screen "eProC - Edición Recetas" 1280x770, template "Template"
   RecipeView "Visor de recetas_1" at 25,54 size 1221x597; Recipe "Pieza"
   TextField "Campo de texto_2" at 43,32 size 125x22; Text 'Edición de Recetas'
   Button "Template_Plantilla_Bouton_12" at 937,715 size 150x53; TextOff 'Ajustes Avanzados SYSTEM'; Authorization "Nivel 2"
      on Press: ActivateScreen("eProC - Avanzado", 0)
   Button "Template_Plantilla_Botón_2" at 128,688 size 150x29; TextOff 'EDICIÓN RECETAS'
   Button "Template_Plantilla_Botón_3" at 129,715 size 150x53; TextOff 'SELECCIÓN RECETAS'
      on Click: ActivateScreen("eProC - Recetas", 0)

screen "HabAlarmas5" 1280x770, template "Template"
   TextField "Campo de texto_1" at 117,85 size 297x18; Text '057 - Falla en Plegador 1 al intentar desactivar fijación'
   TextField "Campo de texto_2" at 117,129 size 357x18; Text '058 - Falla en Plegador 1 al intentar desactivar orden de plegado'
   TextField "Campo de texto_3" at 117,173 size 267x18; Text '059 - Falla en Plegador 1 al intentar subir prensa'
   TextField "Campo de texto_4" at 117,217 size 387x18; Text '060 - Falla en Plegador 1 al intentar bajar primera extensión de prensa'
   TextField "Campo de texto_5" at 117,261 size 297x18; Text '061 - Falla en Plegador 2 al intentar desactivar fijación'
   TextField "Campo de texto_6g" at 117,305 size 357x18; Text '062 - Falla en Plegador 2 al intentar desactivar orden de plegado'
   TextField "Campo de texto_7" at 117,349 size 267x18; Text '063 - Falla en Plegador 2 al intentar subir prensa'
   TextField "Campo de texto_8" at 117,393 size 386x18; Text '064 - Falla en Plegador 2 al intentar subir primera extensión de prensa'
   TextField "Campo de texto_9" at 117,437 size 216x18; Text '065 - Falla al transladar Araña (Avance)'
   TextField "Campo de texto_10" at 117,483 size 135x18; Text '066 - Falla al subir Araña'
   TextField "Campo de texto_11" at 117,525 size 136x18; Text '067 - Falla al bajar Araña'
   TextField "Campo de texto_12" at 117,571 size 135x18; Text '068 - Falla al subir Araña'
   TextField "Campo de texto_13" at 117,613 size 37x18; Text '069 -'
   TextField "Campo de texto_14" at 117,657 size 37x18; Text '070 -'
   Switch "Interruptor_1" at 48,77 size 59x33; TextOff 'SI'; TextOn 'NO'; CaptionText 'Switch'; PictureOff "Check"; PictureOn "UnCheck"
      ProcessValue <- "Desactivar_Falla57"
   Switch "Interruptor_2" at 48,121 size 59x33; TextOff 'SI'; TextOn 'NO'; CaptionText 'Switch'; PictureOff "Check"; PictureOn "UnCheck"
      ProcessValue <- "Desactivar_Falla58"
   Switch "Interruptor_3" at 48,165 size 59x33; TextOff 'SI'; TextOn 'NO'; CaptionText 'Switch'; PictureOff "Check"; PictureOn "UnCheck"
      ProcessValue <- "Desactivar_Falla59"
   Switch "Interruptor_4" at 48,209 size 59x33; TextOff 'SI'; TextOn 'NO'; CaptionText 'Switch'; PictureOff "Check"; PictureOn "UnCheck"
      ProcessValue <- "Desactivar_Falla60"
   Switch "Interruptor_5" at 48,253 size 59x33; TextOff 'SI'; TextOn 'NO'; CaptionText 'Switch'; PictureOff "Check"; PictureOn "UnCheck"
      ProcessValue <- "Desactivar_Falla61"
   Switch "Interruptor_6" at 48,297 size 59x33; TextOff 'SI'; TextOn 'NO'; CaptionText 'Switch'; PictureOff "Check"; PictureOn "UnCheck"
      ProcessValue <- "Desactivar_Falla62"
   Switch "Interruptor_7" at 48,341 size 59x33; TextOff 'SI'; TextOn 'NO'; CaptionText 'Switch'; PictureOff "Check"; PictureOn "UnCheck"
      ProcessValue <- "Desactivar_Falla63"
   Switch "Interruptor_8" at 48,385 size 59x33; TextOff 'SI'; TextOn 'NO'; CaptionText 'Switch'; PictureOff "Check"; PictureOn "UnCheck"
      ProcessValue <- "Desactivar_Falla64"
   Switch "Interruptor_9" at 48,429 size 59x33; TextOff 'SI'; TextOn 'NO'; CaptionText 'Switch'; PictureOff "Check"; PictureOn "UnCheck"
      ProcessValue <- "Desactivar_Falla65"
   Switch "Interruptor_10" at 48,473 size 59x33; TextOff 'SI'; TextOn 'NO'; CaptionText 'Switch'; PictureOff "Check"; PictureOn "UnCheck"
      ProcessValue <- "Desactivar_Falla66"
   Switch "Interruptor_11" at 48,517 size 59x33; TextOff 'SI'; TextOn 'NO'; CaptionText 'Switch'; PictureOff "Check"; PictureOn "UnCheck"
      ProcessValue <- "Desactivar_Falla67"
   Switch "Interruptor_12" at 48,561 size 59x33; TextOff 'SI'; TextOn 'NO'; CaptionText 'Switch'; PictureOff "Check"; PictureOn "UnCheck"
      ProcessValue <- "Desactivar_Falla68"
   Switch "Interruptor_13" at 48,605 size 59x33; TextOff 'SI'; TextOn 'NO'; CaptionText 'Switch'; PictureOff "Check"; PictureOn "UnCheck"
      ProcessValue <- "Desactivar_Falla69"
   Switch "Interruptor_14" at 48,649 size 59x33; TextOff 'SI'; TextOn 'NO'; CaptionText 'Switch'; PictureOff "Check"; PictureOn "UnCheck"
      ProcessValue <- "Desactivar_Falla70"
   TextField "Campo de texto_16" at 664,85 size 37x18; Text '071 -'
   TextField "Campo de texto_17" at 664,129 size 37x18; Text '072 -'
   TextField "Campo de texto_18" at 664,173 size 241x18; Text '073 - Falla al transladar Araña (Retroceder)'
   TextField "Campo de texto_19" at 664,217 size 140x18; Text '074 - Falla al bajar Araña'
   TextField "Campo de texto_20" at 664,261 size 33x18; Text '075 -'
   TextField "Campo de texto_21" at 664,305 size 37x18; Text '076 -'
   TextField "Campo de texto_22" at 664,349 size 392x32; Text '077 - Falla en Plegador 1 al intentar subir segunda extensión de prensa'
   TextField "Campo de texto_23" at 664,393 size 392x32; Text '078 - Falla en Plegador 2 al intentar subir segunda extensión de prensa'
   TextField "Campo de texto_24" at 664,437 size 393x18; Text '079 - Falla en Plegador 1 al intentar bajar segunda extensión de prensa'
   TextField "Campo de texto_25" at 664,483 size 393x18; Text '080 - Falla en Plegador 2 al intentar bajar segunda extensión de prensa'
   TextField "Campo de texto_26" at 664,525 size 219x18; Text '081 - Falla al avanzar ajuste de formado'
   TextField "Campo de texto_27" at 664,571 size 333x18; Text '082 - Falla al subir Bloqueador de Avance en etapa formador'
   TextField "Campo de texto_28" at 664,613 size 206x18; Text '083 - Falla al abrir pinza posicionadora'
   TextField "Campo de texto_29" at 664,657 size 37x18; Text '084 -'
   Switch "Interruptor_15" at 595,77 size 59x33; TextOn 'NO'; TextOff 'SI'; CaptionText 'Switch'; PictureOff "Check"; PictureOn "UnCheck"
      ProcessValue <- "Desactivar_Falla71"
   Switch "Interruptor_16" at 595,121 size 59x33; TextOn 'NO'; TextOff 'SI'; CaptionText 'Switch'; PictureOff "Check"; PictureOn "UnCheck"
      ProcessValue <- "Desactivar_Falla72"
   Switch "Interruptor_17" at 595,165 size 59x33; TextOn 'NO'; TextOff 'SI'; CaptionText 'Switch'; PictureOff "Check"; PictureOn "UnCheck"
      ProcessValue <- "Desactivar_Falla73"
   Switch "Interruptor_18" at 595,209 size 59x33; TextOn 'NO'; TextOff 'SI'; CaptionText 'Switch'; PictureOff "Check"; PictureOn "UnCheck"
      ProcessValue <- "Desactivar_Falla74"
   Switch "Interruptor_19" at 595,253 size 59x33; TextOn 'NO'; TextOff 'SI'; CaptionText 'Switch'; PictureOff "Check"; PictureOn "UnCheck"
      ProcessValue <- "Desactivar_Falla75"
   Switch "Interruptor_20" at 595,297 size 59x33; TextOn 'NO'; TextOff 'SI'; CaptionText 'Switch'; PictureOff "Check"; PictureOn "UnCheck"
      ProcessValue <- "Desactivar_Falla76"
   Switch "Interruptor_21" at 595,341 size 59x33; TextOn 'NO'; TextOff 'SI'; CaptionText 'Switch'; PictureOff "Check"; PictureOn "UnCheck"
      ProcessValue <- "Desactivar_Falla77"
   Switch "Interruptor_22" at 595,385 size 59x33; TextOn 'NO'; TextOff 'SI'; CaptionText 'Switch'; PictureOff "Check"; PictureOn "UnCheck"
      ProcessValue <- "Desactivar_Falla78"
   Switch "Interruptor_23" at 595,429 size 59x33; TextOn 'NO'; TextOff 'SI'; CaptionText 'Switch'; PictureOff "Check"; PictureOn "UnCheck"
      ProcessValue <- "Desactivar_Falla79"
   Switch "Interruptor_24" at 595,473 size 59x33; TextOn 'NO'; TextOff 'SI'; CaptionText 'Switch'; PictureOff "Check"; PictureOn "UnCheck"
      ProcessValue <- "Desactivar_Falla80"
   Switch "Interruptor_25" at 595,517 size 59x33; TextOn 'NO'; TextOff 'SI'; CaptionText 'Switch'; PictureOff "Check"; PictureOn "UnCheck"
      ProcessValue <- "Desactivar_Falla81"
   Switch "Interruptor_26" at 595,561 size 59x33; TextOn 'NO'; TextOff 'SI'; CaptionText 'Switch'; PictureOff "Check"; PictureOn "UnCheck"
      ProcessValue <- "Desactivar_Falla82"
   Switch "Interruptor_27" at 595,605 size 59x33; TextOn 'NO'; TextOff 'SI'; CaptionText 'Switch'; PictureOff "Check"; PictureOn "UnCheck"
      ProcessValue <- "Desactivar_Falla83"
   Switch "Interruptor_28" at 595,649 size 59x33; TextOn 'NO'; TextOff 'SI'; CaptionText 'Switch'; PictureOff "Check"; PictureOn "UnCheck"
      ProcessValue <- "Desactivar_Falla84"
   TextField "Campo de texto_15" at 38,32 size 262x22; Text 'Configuración de habilitación de Alarmas'
   Button "Botón_2" at 1010,33 size 51x51; TextOff '<'
      on Click: ActivateScreen("HabAlarmas3", 0)
   Button "Botón_3" at 1202,33 size 51x51; TextOff '>'
      on Click: ActivateScreen("HabAlarmas7", 0)
   Circle "Círculo_2" at 24,87 size 12x12
      Appearance <- "Alarma 1"
   Circle "Círculo_3" at 25,131 size 12x12
      Appearance <- "Alarma 58"
   Circle "Círculo_4" at 25,175 size 12x12
      Appearance <- "Alarma 59"
   Circle "Círculo_5" at 24,87 size 12x12
      Appearance <- "Alarma 57"
   Circle "Círculo_6" at 25,219 size 12x12
      Appearance <- "Alarma 60"
   Circle "Círculo_7" at 25,263 size 12x12
      Appearance <- "Alarma 61"
   Circle "Círculo_8" at 25,307 size 12x12
      Appearance <- "Alarma 62"
   Circle "Círculo_9" at 25,351 size 12x12
      Appearance <- "Alarma 63"
   Circle "Círculo_10" at 25,395 size 12x12
      Appearance <- "Alarma 64"
   Circle "Círculo_11" at 25,439 size 12x12
      Appearance <- "Alarma 65"
   Circle "Círculo_12" at 25,483 size 12x12
      Appearance <- "Alarma 66"
   Circle "Círculo_13" at 25,527 size 12x12
      Appearance <- "Alarma 67"
   Circle "Círculo_14" at 25,571 size 12x12
      Appearance <- "Alarma 68"
   Circle "Círculo_15" at 25,615 size 12x12
      Appearance <- "Alarma 69"
   Circle "Círculo_16" at 25,659 size 12x12
      Appearance <- "Alarma 70"
   Circle "Círculo_17" at 571,87 size 12x12
      Appearance <- "Alarma 1"
   Circle "Círculo_18" at 572,131 size 12x12
      Appearance <- "Alarma 72"
   Circle "Círculo_19" at 572,175 size 12x12
      Appearance <- "Alarma 73"
   Circle "Círculo_20" at 571,87 size 12x12
      Appearance <- "Alarma 71"
   Circle "Círculo_21" at 572,219 size 12x12
      Appearance <- "Alarma 74"
   Circle "Círculo_22" at 572,263 size 12x12
      Appearance <- "Alarma 75"
   Circle "Círculo_23" at 572,307 size 12x12
      Appearance <- "Alarma 76"
   Circle "Círculo_24" at 572,351 size 12x12
      Appearance <- "Alarma 77"
   Circle "Círculo_26" at 572,395 size 12x12
      Appearance <- "Alarma 78"
   Circle "Círculo_28" at 572,439 size 12x12
      Appearance <- "Alarma 79"
   Circle "Círculo_30" at 572,483 size 12x12
      Appearance <- "Alarma 80"
   Circle "Círculo_32" at 572,527 size 12x12
      Appearance <- "Alarma 81"
   Circle "Círculo_34" at 572,571 size 12x12
      Appearance <- "Alarma 82"
   Circle "Círculo_35" at 572,615 size 12x12
      Appearance <- "Alarma 83"
   Circle "Círculo_36" at 572,659 size 12x12
      Appearance <- "Alarma 84"
   Button "Template_Plantilla_Bouton_0" at 1085,715 size 193x53; TextOff 'ALARMAS / DEFAUT'
      on Press: ActivateScreen("eProC - Alarmas", 0)
   Button "Template_Plantilla_Bouton_2" at 1085,715 size 193x53; TextOff 'ALARMAS / DEFAUT'
      on Press: ActivateScreen("eProC - Alarmas", 0)
      Visibility <- "DB_OP.P_DEFAUT"
   Button "Template_Plantilla_Botón_3" at 1085,688 size 193x29; TextOff 'DESACT. TEMP. ALARMAS'

screen "HabAlarmas1" 1280x770, template "Template"
   TextField "Campo de texto_1" at 117,85 size 394x18; Text '001 - Falla térmica en motor refrigeración de grupo hidráulico Plegadora'
   TextField "Campo de texto_2" at 117,129 size 37x18; Text '002 -'
   TextField "Campo de texto_3" at 117,173 size 317x18; Text '003 - Falla Alimentación Motor Intercambio de Almacenes'
   TextField "Campo de texto_4" at 117,217 size 242x18; Text '004 - Falla en Variador Transporte de Araña'
   TextField "Campo de texto_5" at 117,261 size 221x18; Text '005 - Falla en Variador Transporte Rolos'
   TextField "Campo de texto_6h" at 117,305 size 212x18; Text '006 - Falla en Control Unit Perfiladores'
   TextField "Campo de texto_7" at 117,349 size 323x18; Text '007 - Falla en etapa de Potencia de variadores Perfiladores'
   TextField "Campo de texto_8" at 117,393 size 212x18; Text '008 - Falla presente en CU Plegadores'
   TextField "Campo de texto_9" at 117,437 size 286x18; Text '009 - Falla de seguridad presente en CU Plegadores'
   TextField "Campo de texto_10" at 117,483 size 324x18; Text '010 - Falla térmica en bomba de lubricación de Perfiladores'
   TextField "Campo de texto_11" at 117,525 size 328x18; Text '011 - Falla térmica en grupo hidraulico de freno Perfiladores'
   TextField "Campo de texto_12" at 117,571 size 336x18; Text '012 - Falla térmica en motor Ajuste de ancho de Perfiladores'
   TextField "Campo de texto_13" at 117,613 size 220x18; Text '013 - Falla en Variador Transporte Cinta'
   TextField "Campo de texto_14" at 117,657 size 370x18; Text '014 - Falla térmica en motor ajuste de ancho en etapa de formado'
   Switch "Interruptor_1" at 48,77 size 59x33; TextOff 'SI'; TextOn 'NO'; CaptionText 'Switch'; PictureOff "Check"; PictureOn "UnCheck"
      ProcessValue <- "Desactivar_Falla1"
   Switch "Interruptor_2" at 48,121 size 59x33; TextOff 'SI'; TextOn 'NO'; CaptionText 'Switch'; PictureOff "Check"; PictureOn "UnCheck"
      ProcessValue <- "Desactivar_Falla2"
   Switch "Interruptor_3" at 48,165 size 59x33; TextOff 'SI'; TextOn 'NO'; CaptionText 'Switch'; PictureOff "Check"; PictureOn "UnCheck"
      ProcessValue <- "Desactivar_Falla3"
   Switch "Interruptor_4" at 48,209 size 59x33; TextOff 'SI'; TextOn 'NO'; CaptionText 'Switch'; PictureOff "Check"; PictureOn "UnCheck"
      ProcessValue <- "Desactivar_Falla4"
   Switch "Interruptor_5" at 48,253 size 59x33; TextOff 'SI'; TextOn 'NO'; CaptionText 'Switch'; PictureOff "Check"; PictureOn "UnCheck"
      ProcessValue <- "Desactivar_Falla5"
   Switch "Interruptor_6" at 48,297 size 59x33; TextOff 'SI'; TextOn 'NO'; CaptionText 'Switch'; PictureOff "Check"; PictureOn "UnCheck"
      ProcessValue <- "Desactivar_Falla6"
   Switch "Interruptor_7" at 48,341 size 59x33; TextOff 'SI'; TextOn 'NO'; CaptionText 'Switch'; PictureOff "Check"; PictureOn "UnCheck"
      ProcessValue <- "Desactivar_Falla7"
   Switch "Interruptor_8" at 48,385 size 59x33; TextOff 'SI'; TextOn 'NO'; CaptionText 'Switch'; PictureOff "Check"; PictureOn "UnCheck"
      ProcessValue <- "Desactivar_Falla8"
   Switch "Interruptor_9" at 48,429 size 59x33; TextOff 'SI'; TextOn 'NO'; CaptionText 'Switch'; PictureOff "Check"; PictureOn "UnCheck"
      ProcessValue <- "Desactivar_Falla9"
   Switch "Interruptor_10" at 48,473 size 59x33; TextOff 'SI'; TextOn 'NO'; CaptionText 'Switch'; PictureOff "Check"; PictureOn "UnCheck"
      ProcessValue <- "Desactivar_Falla10"
   Switch "Interruptor_11" at 48,517 size 59x33; TextOff 'SI'; TextOn 'NO'; CaptionText 'Switch'; PictureOff "Check"; PictureOn "UnCheck"
      ProcessValue <- "Desactivar_Falla11"
   Switch "Interruptor_12" at 48,561 size 59x33; TextOff 'SI'; TextOn 'NO'; CaptionText 'Switch'; PictureOff "Check"; PictureOn "UnCheck"
      ProcessValue <- "Desactivar_Falla12"
   Switch "Interruptor_13" at 48,605 size 59x33; TextOff 'SI'; TextOn 'NO'; CaptionText 'Switch'; PictureOff "Check"; PictureOn "UnCheck"
      ProcessValue <- "Desactivar_Falla13"
   Switch "Interruptor_14" at 48,649 size 59x33; TextOff 'SI'; TextOn 'NO'; CaptionText 'Switch'; PictureOff "Check"; PictureOn "UnCheck"
      ProcessValue <- "Desactivar_Falla14"
   Button "Botón_2" at 1010,33 size 51x51; TextOff '<'
   Button "Botón_3" at 1202,33 size 51x51; TextOff '>'
      on Click: ActivateScreen("HabAlarmas3", 0)
   TextField "Campo de texto_16" at 664,85 size 265x18; Text '015 - Falla Rectificador de variadores Plegadores'
   TextField "Campo de texto_17" at 664,129 size 255x18; Text '016 - Falla límite de Seguridad en Plegador 1'
   TextField "Campo de texto_18" at 664,173 size 247x18; Text '017 - Falla límite de Seguridad en Plegador 2'
   TextField "Campo de texto_19" at 664,217 size 305x18; Text '018 - Falla térmica en motor grupo hidráulico Plegadora'
   TextField "Campo de texto_20" at 664,261 size 423x18; Text '019 - Falla térmica en freno de motor ajuste de ancho en etapa de Formado'
   TextField "Campo de texto_21" at 664,305 size 290x18; Text '020 - Falla en presión hidráulica en freno Perfiladores'
   TextField "Campo de texto_22" at 664,349 size 328x18; Text '021 - Falla de excursión en Ajuste de ancho de Perfiladores'
   TextField "Campo de texto_23" at 664,393 size 313x18; Text '022 - Falla de excursión en Ajuste de ancho de Formado'
   TextField "Campo de texto_24" at 664,437 size 208x18; Text '023 - Falla Seguridades de Perímetro'
   TextField "Campo de texto_25" at 664,483 size 37x18; Text '024 -'
   TextField "Campo de texto_26" at 664,525 size 199x18; Text '025 - Falla alimentación de Entradas'
   TextField "Campo de texto_27" at 664,571 size 133x18; Text '026 - Falla de seguridad'
   TextField "Campo de texto_28" at 664,613 size 145x18; Text '027 - Falla presión de Aire'
   TextField "Campo de texto_29" at 664,657 size 226x18; Text '028 - Falla Temperatura Grupo Hidráulico'
   Switch "Interruptor_15" at 595,77 size 59x33; TextOn 'NO'; TextOff 'SI'; CaptionText 'Switch'; PictureOff "Check"; PictureOn "UnCheck"
      ProcessValue <- "Desactivar_Falla15"
   Switch "Interruptor_16" at 595,121 size 59x33; TextOn 'NO'; TextOff 'SI'; CaptionText 'Switch'; PictureOff "Check"; PictureOn "UnCheck"
      ProcessValue <- "Desactivar_Falla16"
   Switch "Interruptor_17" at 595,165 size 59x33; TextOn 'NO'; TextOff 'SI'; CaptionText 'Switch'; PictureOff "Check"; PictureOn "UnCheck"
      ProcessValue <- "Desactivar_Falla17"
   Switch "Interruptor_18" at 595,209 size 59x33; TextOn 'NO'; TextOff 'SI'; CaptionText 'Switch'; PictureOff "Check"; PictureOn "UnCheck"
      ProcessValue <- "Desactivar_Falla18"
   Switch "Interruptor_19" at 595,253 size 59x33; TextOn 'NO'; TextOff 'SI'; CaptionText 'Switch'; PictureOff "Check"; PictureOn "UnCheck"
      ProcessValue <- "Desactivar_Falla19"
   Switch "Interruptor_20" at 595,297 size 59x33; TextOn 'NO'; TextOff 'SI'; CaptionText 'Switch'; PictureOff "Check"; PictureOn "UnCheck"
      ProcessValue <- "Desactivar_Falla20"
   Switch "Interruptor_21" at 595,341 size 59x33; TextOn 'NO'; TextOff 'SI'; CaptionText 'Switch'; PictureOff "Check"; PictureOn "UnCheck"
      ProcessValue <- "Desactivar_Falla21"
   Switch "Interruptor_22" at 595,385 size 59x33; TextOn 'NO'; TextOff 'SI'; CaptionText 'Switch'; PictureOff "Check"; PictureOn "UnCheck"
      ProcessValue <- "Desactivar_Falla22"
   Switch "Interruptor_23" at 595,429 size 59x33; TextOn 'NO'; TextOff 'SI'; CaptionText 'Switch'; PictureOff "Check"; PictureOn "UnCheck"
      ProcessValue <- "Desactivar_Falla23"
   Switch "Interruptor_24" at 595,473 size 59x33; TextOn 'NO'; TextOff 'SI'; CaptionText 'Switch'; PictureOff "Check"; PictureOn "UnCheck"
      ProcessValue <- "Desactivar_Falla24"
   Switch "Interruptor_25" at 595,517 size 59x33; TextOn 'NO'; TextOff 'SI'; CaptionText 'Switch'; PictureOff "Check"; PictureOn "UnCheck"
      ProcessValue <- "Desactivar_Falla25"
   Switch "Interruptor_26" at 595,561 size 59x33; TextOn 'NO'; TextOff 'SI'; CaptionText 'Switch'; PictureOff "Check"; PictureOn "UnCheck"
      ProcessValue <- "Desactivar_Falla26"
   Switch "Interruptor_27" at 595,605 size 59x33; TextOn 'NO'; TextOff 'SI'; CaptionText 'Switch'; PictureOff "Check"; PictureOn "UnCheck"
      ProcessValue <- "Desactivar_Falla27"
   Switch "Interruptor_28" at 595,649 size 59x33; TextOn 'NO'; TextOff 'SI'; CaptionText 'Switch'; PictureOff "Check"; PictureOn "UnCheck"
      ProcessValue <- "Desactivar_Falla28"
   TextField "Campo de texto_15" at 38,32 size 262x22; Text 'Configuración de habilitación de Alarmas'
   Circle "Círculo_2" at 24,87 size 12x12
      Appearance <- "Alarma 1"
   Circle "Círculo_3" at 25,131 size 12x12
      Appearance <- "Alarma 2"
   Circle "Círculo_4" at 25,175 size 12x12
      Appearance <- "Alarma 3"
   Circle "Círculo_5" at 24,87 size 12x12
      Appearance <- "Alarma 1"
   Circle "Círculo_6" at 25,219 size 12x12
      Appearance <- "Alarma 4"
   Circle "Círculo_7" at 25,263 size 12x12
      Appearance <- "Alarma 5"
   Circle "Círculo_8" at 25,307 size 12x12
      Appearance <- "Alarma 6"
   Circle "Círculo_9" at 25,351 size 12x12
      Appearance <- "Alarma 7"
   Circle "Círculo_10" at 25,395 size 12x12
      Appearance <- "Alarma 8"
   Circle "Círculo_11" at 25,439 size 12x12
      Appearance <- "Alarma 9"
   Circle "Círculo_12" at 25,483 size 12x12
      Appearance <- "Alarma 10"
   Circle "Círculo_13" at 25,527 size 12x12
      Appearance <- "Alarma 11"
   Circle "Círculo_14" at 25,571 size 12x12
      Appearance <- "Alarma 12"
   Circle "Círculo_15" at 25,615 size 12x12
      Appearance <- "Alarma 13"
   Circle "Círculo_16" at 25,659 size 12x12
      Appearance <- "Alarma 14"
   Circle "Círculo_17" at 571,87 size 12x12
      Appearance <- "Alarma 1"
   Circle "Círculo_18" at 572,131 size 12x12
      Appearance <- "Alarma 16"
   Circle "Círculo_19" at 572,175 size 12x12
      Appearance <- "Alarma 17"
   Circle "Círculo_20" at 571,87 size 12x12
      Appearance <- "Alarma 15"
   Circle "Círculo_21" at 572,219 size 12x12
      Appearance <- "Alarma 18"
   Circle "Círculo_22" at 572,263 size 12x12
      Appearance <- "Alarma 19"
   Circle "Círculo_23" at 572,307 size 12x12
      Appearance <- "Alarma 20"
   Circle "Círculo_24" at 572,351 size 12x12
      Appearance <- "Alarma 21"
   Circle "Círculo_26" at 572,395 size 12x12
      Appearance <- "Alarma 22"
   Circle "Círculo_28" at 572,439 size 12x12
      Appearance <- "Alarma 23"
   Circle "Círculo_30" at 572,483 size 12x12
      Appearance <- "Alarma 24"
   Circle "Círculo_32" at 572,527 size 12x12
      Appearance <- "Alarma 25"
   Circle "Círculo_34" at 572,571 size 12x12
      Appearance <- "Alarma 26"
   Circle "Círculo_35" at 572,615 size 12x12
      Appearance <- "Alarma 27"
   Circle "Círculo_36" at 572,659 size 12x12
      Appearance <- "Alarma 28"
   Button "Template_Plantilla_Botón_3" at 1085,688 size 193x29; TextOff 'DESACT. TEMP. ALARMAS'
   Button "Template_Plantilla_Bouton_0" at 1085,715 size 193x53; TextOff 'ALARMAS / DEFAUT'
      on Press: ActivateScreen("eProC - Alarmas", 0)
   Button "Template_Plantilla_Bouton_2" at 1085,715 size 193x53; TextOff 'ALARMAS / DEFAUT'
      on Press: ActivateScreen("eProC - Alarmas", 0)
      Visibility <- "DB_OP.P_DEFAUT"

screen "eProC - Tendencia" 1280x770, template "Template"
   IOField "Campo ES_1" at 341,53 size 128x31; FormatPattern 999.99
      ProcessValue <- "Tiempo_Heladera"
      Visibility <- "Hab_Medición"
   IOField "Campo ES_2" at 660,83 size 128x31; FormatPattern 9999.99
      ProcessValue <- "HeladerasxHora"
      Visibility <- "Hab_Medición"
   IOField "Campo ES_3" at 660,51 size 128x31; FormatPattern 9999.99
      ProcessValue <- "HeladerasxMin"
      Visibility <- "Hab_Medición"
   TextField "Campo de texto_16" at 728,54 size 114x22; Text 'Heladeras x Min.'
      Visibility <- "Hab_Medición"
   TextField "Campo de texto_17" at 728,86 size 118x22; Text 'Heladeras x Hora'
      Visibility <- "Hab_Medición"
   IOField "Campo ES_4" at 341,85 size 128x31; FormatPattern 999.99
      ProcessValue <- "Tiempo_Heladera_Prom"
      Visibility <- "Hab_Medición"
   TextField "Campo de texto_19" at 402,88 size 143x22; Text 'Segundos x Heladera'
      Visibility <- "Hab_Medición"
   TextField "Campo de texto_20" at 402,56 size 143x22; Text 'Segundos x Heladera'
      Visibility <- "Hab_Medición"
   TextField "Campo de texto_21" at 227,56 size 107x22; Text 'Última Heladera'
      Visibility <- "Hab_Medición"
   TextField "Campo de texto_22" at 162,88 size 174x22; Text 'Tendencia (10 Heladeras)'
      Visibility <- "Hab_Medición"
   TrendView "Visualización de curvas_1" at 90,192 size 1062x427

screen "HabAlarmas3" 1280x770, template "Template"
   TextField "Campo de texto_1" at 117,85 size 248x18; Text '029 - Falla Seguridad Barrera en Descargador'
   TextField "Campo de texto_2" at 117,129 size 184x18; Text '030 - Falla Cubierta de Perfilador'
   TextField "Campo de texto_3" at 117,173 size 239x18; Text '031 - Falla de Atasco de pieza en Perfilador'
   TextField "Campo de texto_4" at 117,217 size 37x18; Text '032 -'
   TextField "Campo de texto_5" at 117,261 size 225x18; Text '033 - Falla avance de pinza en Plegadora'
   TextField "Campo de texto_6ñ" at 117,305 size 207x18; Text '034 - Falla al bajar pinza en Plegadora'
   TextField "Campo de texto_7" at 117,349 size 204x18; Text '035 - Falla al abrir pinza en Plegadora'
   TextField "Campo de texto_8" at 117,393 size 301x18; Text '036 - Falla al activar alineacion X de Pieza en Plegadora'
   TextField "Campo de texto_9" at 117,437 size 302x18; Text '037 - Falla al activar alineacion Y de Pieza en Plegadora'
   TextField "Campo de texto_10" at 117,483 size 321x18; Text '038 - Falla al desactivar alineacion Y de Pieza en Plegadora'
   TextField "Campo de texto_11" at 117,525 size 33x18; Text '039 -'
   TextField "Campo de texto_12" at 117,571 size 37x18; Text '040 -'
   TextField "Campo de texto_13" at 117,613 size 239x18; Text '041 - Falla retroceso de pinza en Plegadora'
   TextField "Campo de texto_14" at 117,657 size 206x18; Text '042 - Falla al subir pinza en Plegadora'
   Switch "Interruptor_1" at 48,77 size 59x33; TextOff 'SI'; TextOn 'NO'; CaptionText 'Switch'; PictureOff "Check"; PictureOn "UnCheck"
      ProcessValue <- "Desactivar_Falla29"
   Switch "Interruptor_2" at 48,121 size 59x33; TextOff 'SI'; TextOn 'NO'; CaptionText 'Switch'; PictureOff "Check"; PictureOn "UnCheck"
      ProcessValue <- "Desactivar_Falla30"
   Switch "Interruptor_3" at 48,165 size 59x33; TextOff 'SI'; TextOn 'NO'; CaptionText 'Switch'; PictureOff "Check"; PictureOn "UnCheck"
      ProcessValue <- "Desactivar_Falla31"
   Switch "Interruptor_4" at 48,209 size 59x33; TextOff 'SI'; TextOn 'NO'; CaptionText 'Switch'; PictureOff "Check"; PictureOn "UnCheck"
      ProcessValue <- "Desactivar_Falla32"
   Switch "Interruptor_5" at 48,253 size 59x33; TextOff 'SI'; TextOn 'NO'; CaptionText 'Switch'; PictureOff "Check"; PictureOn "UnCheck"
      ProcessValue <- "Desactivar_Falla33"
   Switch "Interruptor_6" at 48,297 size 59x33; TextOff 'SI'; TextOn 'NO'; CaptionText 'Switch'; PictureOff "Check"; PictureOn "UnCheck"
      ProcessValue <- "Desactivar_Falla34"
   Switch "Interruptor_7" at 48,341 size 59x33; TextOff 'SI'; TextOn 'NO'; CaptionText 'Switch'; PictureOff "Check"; PictureOn "UnCheck"
      ProcessValue <- "Desactivar_Falla35"
   Switch "Interruptor_8" at 48,385 size 59x33; TextOff 'SI'; TextOn 'NO'; CaptionText 'Switch'; PictureOff "Check"; PictureOn "UnCheck"
      ProcessValue <- "Desactivar_Falla36"
   Switch "Interruptor_9" at 48,429 size 59x33; TextOff 'SI'; TextOn 'NO'; CaptionText 'Switch'; PictureOff "Check"; PictureOn "UnCheck"
      ProcessValue <- "Desactivar_Falla37"
   Switch "Interruptor_10" at 48,473 size 59x33; TextOff 'SI'; TextOn 'NO'; CaptionText 'Switch'; PictureOff "Check"; PictureOn "UnCheck"
      ProcessValue <- "Desactivar_Falla38"
   Switch "Interruptor_11" at 48,517 size 59x33; TextOff 'SI'; TextOn 'NO'; CaptionText 'Switch'; PictureOff "Check"; PictureOn "UnCheck"
      ProcessValue <- "Desactivar_Falla39"
   Switch "Interruptor_12" at 48,561 size 59x33; TextOff 'SI'; TextOn 'NO'; CaptionText 'Switch'; PictureOff "Check"; PictureOn "UnCheck"
      ProcessValue <- "Desactivar_Falla40"
   Switch "Interruptor_13" at 48,605 size 59x33; TextOff 'SI'; TextOn 'NO'; CaptionText 'Switch'; PictureOff "Check"; PictureOn "UnCheck"
      ProcessValue <- "Desactivar_Falla41"
   Switch "Interruptor_14" at 48,649 size 59x33; TextOff 'SI'; TextOn 'NO'; CaptionText 'Switch'; PictureOff "Check"; PictureOn "UnCheck"
      ProcessValue <- "Desactivar_Falla42"
   TextField "Campo de texto_16" at 664,85 size 212x18; Text '043 - Falla al cerrar pinza en Plegadora'
   TextField "Campo de texto_17" at 664,129 size 320x18; Text '044 - Falla al desactivar alineacion X de Pieza en Plegadora'
   TextField "Campo de texto_18" at 664,173 size 321x18; Text '045 - Falla al desactivar alineacion Y de Pieza en Plegadora'
   TextField "Campo de texto_19" at 664,217 size 218x18; Text '046 - Falla al Bajar cepillos en Plegadora'
   TextField "Campo de texto_20" at 664,261 size 37x18; Text '047 -'
   TextField "Campo de texto_21" at 664,305 size 37x18; Text '048 -'
   TextField "Campo de texto_22" at 664,349 size 278x18; Text '049 - Falla en Plegador 1 al intentar activar fijación'
   TextField "Campo de texto_23" at 664,393 size 285x18; Text '050 - Falla en Plegador 1 al intentar realizar plegado'
   TextField "Campo de texto_24" at 664,437 size 268x18; Text '051 - Falla en Plegador 1 al intentar bajar prensa'
   TextField "Campo de texto_25" at 664,483 size 386x18; Text '052 - Falla en Plegador 1 al intentar subir primera extensión de prensa'
   TextField "Campo de texto_26" at 664,525 size 278x18; Text '053 - Falla en Plegador 2 al intentar activar fijación'
   TextField "Campo de texto_27" at 664,571 size 285x18; Text '054 - Falla en Plegador 2 al intentar realizar plegado'
   TextField "Campo de texto_28" at 664,613 size 268x18; Text '055 - Falla en Plegador 2 al intentar bajar prensa'
   TextField "Campo de texto_29" at 664,657 size 387x18; Text '056 - Falla en Plegador 2 al intentar bajar primera extensión de prensa'
   Switch "Interruptor_15" at 595,77 size 59x33; TextOn 'NO'; TextOff 'SI'; CaptionText 'Switch'; PictureOff "Check"; PictureOn "UnCheck"
      ProcessValue <- "Desactivar_Falla43"
   Switch "Interruptor_16" at 595,121 size 59x33; TextOn 'NO'; TextOff 'SI'; CaptionText 'Switch'; PictureOff "Check"; PictureOn "UnCheck"
      ProcessValue <- "Desactivar_Falla44"
   Switch "Interruptor_17" at 595,165 size 59x33; TextOn 'NO'; TextOff 'SI'; CaptionText 'Switch'; PictureOff "Check"; PictureOn "UnCheck"
      ProcessValue <- "Desactivar_Falla45"
   Switch "Interruptor_18" at 595,209 size 59x33; TextOn 'NO'; TextOff 'SI'; CaptionText 'Switch'; PictureOff "Check"; PictureOn "UnCheck"
      ProcessValue <- "Desactivar_Falla46"
   Switch "Interruptor_19" at 595,253 size 59x33; TextOn 'NO'; TextOff 'SI'; CaptionText 'Switch'; PictureOff "Check"; PictureOn "UnCheck"
      ProcessValue <- "Desactivar_Falla47"
   Switch "Interruptor_20" at 595,297 size 59x33; TextOn 'NO'; TextOff 'SI'; CaptionText 'Switch'; PictureOff "Check"; PictureOn "UnCheck"
      ProcessValue <- "Desactivar_Falla48"
   Switch "Interruptor_21" at 595,341 size 59x33; TextOn 'NO'; TextOff 'SI'; CaptionText 'Switch'; PictureOff "Check"; PictureOn "UnCheck"
      ProcessValue <- "Desactivar_Falla49"
   Switch "Interruptor_22" at 595,385 size 59x33; TextOn 'NO'; TextOff 'SI'; CaptionText 'Switch'; PictureOff "Check"; PictureOn "UnCheck"
      ProcessValue <- "Desactivar_Falla50"
   Switch "Interruptor_23" at 595,429 size 59x33; TextOn 'NO'; TextOff 'SI'; CaptionText 'Switch'; PictureOff "Check"; PictureOn "UnCheck"
      ProcessValue <- "Desactivar_Falla51"
   Switch "Interruptor_24" at 595,473 size 59x33; TextOn 'NO'; TextOff 'SI'; CaptionText 'Switch'; PictureOff "Check"; PictureOn "UnCheck"
      ProcessValue <- "Desactivar_Falla52"
   Switch "Interruptor_25" at 595,517 size 59x33; TextOn 'NO'; TextOff 'SI'; CaptionText 'Switch'; PictureOff "Check"; PictureOn "UnCheck"
      ProcessValue <- "Desactivar_Falla53"
   Switch "Interruptor_26" at 595,561 size 59x33; TextOn 'NO'; TextOff 'SI'; CaptionText 'Switch'; PictureOff "Check"; PictureOn "UnCheck"
      ProcessValue <- "Desactivar_Falla54"
   Switch "Interruptor_27" at 595,605 size 59x33; TextOn 'NO'; TextOff 'SI'; CaptionText 'Switch'; PictureOff "Check"; PictureOn "UnCheck"
      ProcessValue <- "Desactivar_Falla55"
   Switch "Interruptor_28" at 595,649 size 59x33; TextOn 'NO'; TextOff 'SI'; CaptionText 'Switch'; PictureOff "Check"; PictureOn "UnCheck"
      ProcessValue <- "Desactivar_Falla56"
   TextField "Campo de texto_15" at 38,32 size 262x22; Text 'Configuración de habilitación de Alarmas'
   Button "Botón_2" at 1010,33 size 51x51; TextOff '<'
      on Click: ActivateScreen("HabAlarmas1", 0)
   Button "Botón_3" at 1202,33 size 51x51; TextOff '>'
      on Click: ActivateScreen("HabAlarmas5", 0)
   Circle "Círculo_2" at 24,87 size 12x12
      Appearance <- "Alarma 1"
   Circle "Círculo_3" at 25,131 size 12x12
      Appearance <- "Alarma 30"
   Circle "Círculo_4" at 25,175 size 12x12
      Appearance <- "Alarma 31"
   Circle "Círculo_5" at 24,87 size 12x12
      Appearance <- "Alarma 29"
   Circle "Círculo_6" at 25,219 size 12x12
      Appearance <- "Alarma 32"
   Circle "Círculo_7" at 25,263 size 12x12
      Appearance <- "Alarma 33"
   Circle "Círculo_8" at 25,307 size 12x12
      Appearance <- "Alarma 34"
   Circle "Círculo_9" at 25,351 size 12x12
      Appearance <- "Alarma 35"
   Circle "Círculo_10" at 25,395 size 12x12
      Appearance <- "Alarma 36"
   Circle "Círculo_11" at 25,439 size 12x12
      Appearance <- "Alarma 37"
   Circle "Círculo_12" at 25,483 size 12x12
      Appearance <- "Alarma 38"
   Circle "Círculo_13" at 25,527 size 12x12
      Appearance <- "Alarma 39"
   Circle "Círculo_14" at 25,571 size 12x12
      Appearance <- "Alarma 40"
   Circle "Círculo_15" at 25,615 size 12x12
      Appearance <- "Alarma 41"
   Circle "Círculo_16" at 25,659 size 12x12
      Appearance <- "Alarma 42"
   Circle "Círculo_17" at 571,87 size 12x12
      Appearance <- "Alarma 1"
   Circle "Círculo_18" at 572,131 size 12x12
      Appearance <- "Alarma 44"
   Circle "Círculo_19" at 572,175 size 12x12
      Appearance <- "Alarma 45"
   Circle "Círculo_20" at 571,87 size 12x12
      Appearance <- "Alarma 43"
   Circle "Círculo_21" at 572,219 size 12x12
      Appearance <- "Alarma 46"
   Circle "Círculo_22" at 572,263 size 12x12
      Appearance <- "Alarma 47"
   Circle "Círculo_23" at 572,307 size 12x12
      Appearance <- "Alarma 48"
   Circle "Círculo_24" at 572,351 size 12x12
      Appearance <- "Alarma 49"
   Circle "Círculo_26" at 572,395 size 12x12
      Appearance <- "Alarma 50"
   Circle "Círculo_28" at 572,439 size 12x12
      Appearance <- "Alarma 51"
   Circle "Círculo_30" at 572,483 size 12x12
      Appearance <- "Alarma 52"
   Circle "Círculo_32" at 572,527 size 12x12
      Appearance <- "Alarma 53"
   Circle "Círculo_34" at 572,571 size 12x12
      Appearance <- "Alarma 54"
   Circle "Círculo_35" at 572,615 size 12x12
      Appearance <- "Alarma 55"
   Circle "Círculo_36" at 572,659 size 12x12
      Appearance <- "Alarma 56"
   Button "Template_Plantilla_Bouton_0" at 1085,715 size 193x53; TextOff 'ALARMAS / DEFAUT'
      on Press: ActivateScreen("eProC - Alarmas", 0)
   Button "Template_Plantilla_Bouton_2" at 1085,715 size 193x53; TextOff 'ALARMAS / DEFAUT'
      on Press: ActivateScreen("eProC - Alarmas", 0)
      Visibility <- "DB_OP.P_DEFAUT"
   Button "Template_Plantilla_Botón_3" at 1085,688 size 193x29; TextOff 'DESACT. TEMP. ALARMAS'

screen "eProC - Seguimiento Datos" 1280x770, template "Template"
   TextField "Campo de texto_9" at 150,77 size 35x18; Text 'Araña'
   TextField "Campo de texto_10" at 327,77 size 32x18; Text 'Rolos'
   TextField "Campo de texto_11" at 501,77 size 54x18; Text 'Perfilador'
   TextField "Campo de texto_12" at 850,77 size 31x18; Text 'Pinza'
   TextField "Campo de texto_13" at 1029,77 size 57x18; Text 'Plegadora'
   TextField "Campo de texto_16" at 150,130 size 12x18; Text 'A'
   IOField "Champ E/S_8" at 171,127 size 54x25; FormatPattern 9999999
      Appearance <- "Araña\Araña.PresenciaPieza"
      ProcessValue <- "Araña\Araña.A"
   IOField "Champ E/S_9" at 171,147 size 54x25; FormatPattern 9999999
      Appearance <- "Araña\Araña.PresenciaPieza"
      ProcessValue <- "Araña\Araña.B"
   IOField "Champ E/S_10" at 171,168 size 54x24; FormatPattern 9999999
      Appearance <- "Araña\Araña.PresenciaPieza"
      ProcessValue <- "Araña\Araña.C"
   IOField "Champ E/S_11" at 171,187 size 54x25; FormatPattern 9999999
      Appearance <- "Araña\Araña.PresenciaPieza"
      ProcessValue <- "Araña\Araña.D"
   TextField "Campo de texto_17" at 151,148 size 11x18; Text 'B'
   TextField "Campo de texto_18" at 151,168 size 11x18; Text 'C'
   TextField "Campo de texto_19" at 151,188 size 12x18; Text 'D'
   TextField "Campo de texto_20" at 327,131 size 12x18; Text 'A'
   IOField "Champ E/S_12" at 346,127 size 54x25; FormatPattern 9999999
      Appearance <- "Rolos\Rolos.PresenciaPieza"
      ProcessValue <- "Rolos\Rolos.A"
   IOField "Champ E/S_13" at 346,147 size 54x25; FormatPattern 9999999
      Appearance <- "Rolos\Rolos.PresenciaPieza"
      ProcessValue <- "Rolos\Rolos.B"
   IOField "Champ E/S_14" at 346,168 size 54x24; FormatPattern 9999999
      Appearance <- "Rolos\Rolos.PresenciaPieza"
      ProcessValue <- "Rolos\Rolos.C"
   IOField "Champ E/S_15" at 346,187 size 54x25; FormatPattern 9999999
      Appearance <- "Rolos\Rolos.PresenciaPieza"
      ProcessValue <- "Rolos\Rolos.D"
   TextField "Campo de texto_21" at 327,149 size 11x18; Text 'B'
   TextField "Campo de texto_22" at 327,169 size 11x18; Text 'C'
   TextField "Campo de texto_23" at 327,189 size 12x18; Text 'D'
   TextField "Campo de texto_24" at 501,131 size 12x18; Text 'A'
   IOField "Champ E/S_16" at 524,127 size 53x25; FormatPattern 9999999
      Appearance <- "Perfiladores\Perfilador.PresenciaPieza"
      ProcessValue <- "Perfiladores\Perfilador.A"
   IOField "Champ E/S_17" at 524,147 size 53x25; FormatPattern 9999999
      Appearance <- "Perfiladores\Perfilador.PresenciaPieza"
      ProcessValue <- "Perfiladores\Perfilador.B"
   IOField "Champ E/S_18" at 524,168 size 53x24; FormatPattern 9999999
      Appearance <- "Perfiladores\Perfilador.PresenciaPieza"
      ProcessValue <- "Perfiladores\Perfilador.C"
   IOField "Champ E/S_19" at 524,187 size 53x25; FormatPattern 9999999
      Appearance <- "Perfiladores\Perfilador.PresenciaPieza"
      ProcessValue <- "Perfiladores\Perfilador.D"
   TextField "Campo de texto_25" at 503,149 size 11x18; Text 'B'
   TextField "Campo de texto_26" at 503,169 size 11x18; Text 'C'
   TextField "Campo de texto_27" at 503,189 size 12x18; Text 'D'
   TextField "Campo de texto_28" at 850,131 size 12x18; Text 'A'
   IOField "Champ E/S_20" at 875,127 size 53x25; FormatPattern 9999999
      Appearance <- "Pinza\Pinza.PresenciaPieza"
      ProcessValue <- "Pinza\Pinza.A"
   IOField "Champ E/S_21" at 875,147 size 53x25; FormatPattern 9999999
      Appearance <- "Pinza\Pinza.PresenciaPieza"
      ProcessValue <- "Pinza\Pinza.B"
   IOField "Champ E/S_22" at 875,168 size 53x24; FormatPattern 9999999
      Appearance <- "Pinza\Pinza.PresenciaPieza"
      ProcessValue <- "Pinza\Pinza.C"
   IOField "Champ E/S_23" at 875,187 size 53x25; FormatPattern 9999999
      Appearance <- "Pinza\Pinza.PresenciaPieza"
      ProcessValue <- "Pinza\Pinza.D"
   TextField "Campo de texto_29" at 850,149 size 11x18; Text 'B'
   TextField "Campo de texto_30" at 850,169 size 11x18; Text 'C'
   TextField "Campo de texto_31" at 850,189 size 12x18; Text 'D'
   TextField "Campo de texto_32" at 1029,131 size 12x18; Text 'A'
   IOField "Champ E/S_24" at 1050,127 size 53x25; FormatPattern 9999999
      Appearance <- "Plegadora\Plegadora.PresenciaPieza"
      ProcessValue <- "Plegadora\Plegadora.A"
   IOField "Champ E/S_25" at 1050,147 size 53x25; FormatPattern 9999999
      Appearance <- "Plegadora\Plegadora.PresenciaPieza"
      ProcessValue <- "Plegadora\Plegadora.B"
   IOField "Champ E/S_26" at 1050,168 size 53x24; FormatPattern 9999999
      Appearance <- "Plegadora\Plegadora.PresenciaPieza"
      ProcessValue <- "Plegadora\Plegadora.C"
   IOField "Champ E/S_27" at 1050,187 size 53x25; FormatPattern 9999999
      Appearance <- "Plegadora\Plegadora.PresenciaPieza"
      ProcessValue <- "Plegadora\Plegadora.D"
   TextField "Campo de texto_33" at 1029,149 size 11x18; Text 'B'
   TextField "Campo de texto_34" at 1029,169 size 11x18; Text 'C'
   TextField "Campo de texto_35" at 1029,189 size 12x18; Text 'D'
   Button "Botón_8" at 499,38 size 80x36; TextOff 'Borrar'; PictureOff "Borrar Pulsador"
      on Click: ResetBit("Perfiladores\Perfilador.PresenciaPieza")
      Visibility <- "Perfiladores\Perfilador.PresenciaPieza"
   Button "Botón_9" at 325,38 size 80x36; TextOff 'Borrar'; PictureOff "Borrar Pulsador"
      on Click: ResetBit("Rolos\Rolos.PresenciaPieza")
      Visibility <- "Rolos\Rolos.PresenciaPieza"
   Button "Botón_10" at 148,38 size 80x36; TextOff 'Borrar'; PictureOff "Borrar Pulsador"
      on Click: ResetBit("Araña\Araña.PresenciaPieza")
      Visibility <- "Araña\Araña.PresenciaPieza"
   TextField "Campo de texto_113" at 677,77 size 31x18; Text 'Cinta'
   TextField "Campo de texto_114" at 677,131 size 12x18; Text 'A'
   IOField "Champ E/S_106" at 700,127 size 53x25; FormatPattern 9999999
      Appearance <- "Cinta\Cinta.PresenciaPieza"
      ProcessValue <- "Cinta\Cinta.A"
   IOField "Champ E/S_107" at 700,147 size 53x25; FormatPattern 9999999
      Appearance <- "Cinta\Cinta.PresenciaPieza"
      ProcessValue <- "Cinta\Cinta.B"
   IOField "Champ E/S_108" at 700,168 size 53x24; FormatPattern 9999999
      Appearance <- "Cinta\Cinta.PresenciaPieza"
      ProcessValue <- "Cinta\Cinta.C"
   IOField "Champ E/S_109" at 700,187 size 53x25; FormatPattern 9999999
      Appearance <- "Cinta\Cinta.PresenciaPieza"
      ProcessValue <- "Cinta\Cinta.D"
   TextField "Campo de texto_115" at 677,149 size 11x18; Text 'B'
   TextField "Campo de texto_116" at 677,169 size 11x18; Text 'C'
   TextField "Campo de texto_117" at 677,189 size 12x18; Text 'D'
   Button "Botón_14" at 675,38 size 80x36; TextOff 'Borrar'; PictureOff "Borrar Pulsador"
      on Click: ResetBit("Cinta\Cinta.PresenciaPieza")
      Visibility <- "Cinta\Cinta.PresenciaPieza"
   Button "Botón_15" at 850,38 size 80x36; TextOff 'Borrar'; PictureOff "Borrar Pulsador"
      on Click: ResetBit("Pinza\Pinza.PresenciaPieza")
      Visibility <- "Pinza\Pinza.PresenciaPieza"
   Button "Botón_16" at 1025,38 size 80x36; TextOff 'Borrar'; PictureOff "Borrar Pulsador"
      on Click: ResetBit("Plegadora\Plegadora.PresenciaPieza")
      Visibility <- "Plegadora\Plegadora.PresenciaPieza"
   GraphicView "Visor de gráficos_2" at 273,77 size 29x29; Picture "Gráfico_4"
   GraphicView "Visor de gráficos_1" at 446,77 size 29x29; Picture "Gráfico_4"
   GraphicView "Visor de gráficos_3" at 623,77 size 29x29; Picture "Gráfico_4"
   GraphicView "Visor de gráficos_4" at 796,77 size 29x29; Picture "Gráfico_4"
   GraphicView "Visor de gráficos_5" at 971,77 size 29x29; Picture "Gráfico_4"
   TextField "Campo de texto_1" at 72,425 size 54x29; Text 'Pinza'
   TextField "Campo de texto_2" at 229,507 size 54x18; Text 'Solicitada'
   TextField "Campo de texto_49" at 142,529 size 60x18; Text 'Recepción'
   IOField "Champ E/S_1" at 221,525 size 85x25; FormatPattern s9999999999
      ProcessValue <- "Pos_Recepcion"
      Appearance <- "Pinza\Pinza.PresenciaPieza"
   IOField "Champ E/S_2" at 221,545 size 85x25; FormatPattern s9999999999
      ProcessValue <- "Pos_E1H1"
      Appearance <- "Pinza\Pinza.PresenciaPieza"
   IOField "Champ E/S_3" at 221,566 size 85x24; FormatPattern s9999999999
      ProcessValue <- "Pos_E1H2"
      Appearance <- "Pinza\Pinza.PresenciaPieza"
   IOField "Champ E/S_4" at 221,585 size 85x25; FormatPattern s9999999999
      ProcessValue <- "Pos_E2H1"
      Appearance <- "Pinza\Pinza.PresenciaPieza"
   TextField "Campo de texto_50" at 142,547 size 33x18; Text 'E1H1'
   TextField "Campo de texto_51" at 142,567 size 33x18; Text 'E1H2'
   TextField "Campo de texto_52" at 142,587 size 33x18; Text 'E2H1'
   TextField "Campo de texto_53" at 313,507 size 57x18; Text 'Alcanzada'
   IOField "Champ E/S_5" at 305,525 size 85x25; FormatPattern s9999999999
      ProcessValue <- "Pos_Recepcion(3)"
      Appearance <- "Pinza\Pinza.PresenciaPieza"
   IOField "Champ E/S_6" at 305,545 size 85x25; FormatPattern s9999999999
      ProcessValue <- "Pos_E1H1(3)"
      Appearance <- "Pinza\Pinza.PresenciaPieza"
   IOField "Champ E/S_7" at 305,566 size 85x24; FormatPattern s9999999999
      ProcessValue <- "Pos_E1H2(3)"
      Appearance <- "Pinza\Pinza.PresenciaPieza"
   IOField "Champ E/S_28" at 305,585 size 85x25; FormatPattern s9999999999
      ProcessValue <- "Pos_E2H1(3)"
      Appearance <- "Pinza\Pinza.PresenciaPieza"
   TextField "Campo de texto_65" at 615,507 size 54x18; Text 'Solicitada'
   IOField "Champ E/S_57" at 608,525 size 85x25; FormatPattern s9999999999
      ProcessValue <- "Pos_Recepcion(1)"
      Appearance <- "Pinza\Pinza.PresenciaPieza"
   IOField "Champ E/S_58" at 608,545 size 85x25; FormatPattern s9999999999
      ProcessValue <- "Pos_E1H1(1)"
      Appearance <- "Pinza\Pinza.PresenciaPieza"
   IOField "Champ E/S_59" at 608,566 size 85x24; FormatPattern s9999999999
      ProcessValue <- "Pos_E1H2(1)"
      Appearance <- "Pinza\Pinza.PresenciaPieza"
   IOField "Champ E/S_60" at 608,585 size 85x25; FormatPattern s9999999999
      ProcessValue <- "Pos_E2H1(1)"
      Appearance <- "Pinza\Pinza.PresenciaPieza"
   TextField "Campo de texto_78" at 697,507 size 57x18; Text 'Alcanzada'
   IOField "Champ E/S_69" at 690,525 size 85x25; FormatPattern s9999999999
      ProcessValue <- "Pos_Recepcion(4)"
      Appearance <- "Pinza\Pinza.PresenciaPieza"
   IOField "Champ E/S_70" at 690,545 size 85x25; FormatPattern s9999999999
      ProcessValue <- "Pos_E1H1(4)"
      Appearance <- "Pinza\Pinza.PresenciaPieza"
   IOField "Champ E/S_71" at 690,566 size 85x24; FormatPattern s9999999999
      ProcessValue <- "Pos_E1H2(4)"
      Appearance <- "Pinza\Pinza.PresenciaPieza"
   IOField "Champ E/S_72" at 690,585 size 85x25; FormatPattern s9999999999
      ProcessValue <- "Pos_E2H1(4)"
      Appearance <- "Pinza\Pinza.PresenciaPieza"
   TextField "Campo de texto_91" at 1003,507 size 54x18; Text 'Solicitada'
   IOField "Champ E/S_81" at 995,525 size 85x25; FormatPattern s9999999999
      ProcessValue <- "Pos_Recepcion(2)"
      Appearance <- "Pinza\Pinza.PresenciaPieza"
   IOField "Champ E/S_82" at 995,545 size 85x25; FormatPattern s9999999999
      ProcessValue <- "Pos_E1H1(2)"
      Appearance <- "Pinza\Pinza.PresenciaPieza"
   IOField "Champ E/S_83" at 995,566 size 85x24; FormatPattern s9999999999
      ProcessValue <- "Pos_E1H2(2)"
      Appearance <- "Pinza\Pinza.PresenciaPieza"
   IOField "Champ E/S_84" at 995,585 size 85x25; FormatPattern s9999999999
      ProcessValue <- "Pos_E2H1(2)"
      Appearance <- "Pinza\Pinza.PresenciaPieza"
   TextField "Campo de texto_104" at 1085,507 size 57x18; Text 'Alcanzada'
   IOField "Champ E/S_93" at 1077,525 size 85x25; FormatPattern s9999999999
      ProcessValue <- "Pos_Recepcion(5)"
      Appearance <- "Pinza\Pinza.PresenciaPieza"
   IOField "Champ E/S_94" at 1077,545 size 85x25; FormatPattern s9999999999
      ProcessValue <- "Pos_E1H1(5)"
      Appearance <- "Pinza\Pinza.PresenciaPieza"
   IOField "Champ E/S_95" at 1077,566 size 85x24; FormatPattern s9999999999
      ProcessValue <- "Pos_E1H2(5)"
      Appearance <- "Pinza\Pinza.PresenciaPieza"
   IOField "Champ E/S_96" at 1077,585 size 85x25; FormatPattern s9999999999
      ProcessValue <- "Pos_E2H1(5)"
      Appearance <- "Pinza\Pinza.PresenciaPieza"
   TextField "Campo de texto_55" at 533,529 size 60x18; Text 'Recepción'
   TextField "Campo de texto_56" at 533,547 size 33x18; Text 'E1H1'
   TextField "Campo de texto_57" at 533,567 size 33x18; Text 'E1H2'
   TextField "Campo de texto_58" at 533,587 size 33x18; Text 'E2H1'
   TextField "Campo de texto_59" at 916,529 size 60x18; Text 'Recepción'
   TextField "Campo de texto_60" at 916,547 size 33x18; Text 'E1H1'
   TextField "Campo de texto_61" at 916,567 size 33x18; Text 'E1H2'
   TextField "Campo de texto_62" at 916,587 size 33x18; Text 'E2H1'
   TextField "Campo de texto_63" at 231,488 size 128x18; Text 'Posición pieza anterior:'
   TextField "Campo de texto_64" at 616,488 size 139x18; Text 'Posición pieza anterior 2:'
   TextField "Campo de texto_66" at 1002,488 size 139x18; Text 'Posición pieza anterior 3:'
   Button "Template_Plantilla_Botón_3" at 275,715 size 150x53; TextOff 'SEGUIMIENTO DE DATOS'
      on Click: ActivateScreen("eProC - Recetas", 0)
   Button "Template_Plantilla_Bouton_2" at 1085,715 size 193x53; TextOff 'ALARMAS / DEFAUT'
      on Press: ActivateScreen("eProC - Alarmas", 0)
      Visibility <- "DB_OP.P_DEFAUT"
   TextField "Campo de texto_118" at 503,210 size 17x18; Text 'F1'
   IOField "Champ E/S_110" at 527,207 size 51x25; FormatPattern s999999
      Appearance <- "Perfiladores\Perfilador.PresenciaPieza"
      ProcessValue <- "Perfiladores\Perfilador.F1"
   IOField "Champ E/S_111" at 527,227 size 51x25; FormatPattern s999999
      Appearance <- "Perfiladores\Perfilador.PresenciaPieza"
      ProcessValue <- "Perfiladores\Perfilador.F2"
   IOField "Champ E/S_112" at 527,248 size 51x24; FormatPattern s999999
      Appearance <- "Perfiladores\Perfilador.PresenciaPieza"
      ProcessValue <- "Perfiladores\Perfilador.F3"
   IOField "Champ E/S_113" at 527,267 size 51x25; FormatPattern s999999
      Appearance <- "Perfiladores\Perfilador.PresenciaPieza"
      ProcessValue <- "Perfiladores\Perfilador.F4"
   TextField "Campo de texto_119" at 503,229 size 17x18; Text 'F2'
   TextField "Campo de texto_120" at 503,249 size 17x18; Text 'F3'
   TextField "Campo de texto_121" at 503,269 size 17x18; Text 'F4'
   TextField "Campo de texto_122" at 503,290 size 35x18; Text 'PL1-1'
   IOField "Champ E/S_114" at 543,287 size 51x25; FormatPattern s999999
      Appearance <- "Perfiladores\Perfilador.PresenciaPieza"